
   // Not- Aus Taster Farbe 01 -- DB810.DBX67.5
   //    UN    "NA_SchrankFarbe"
   //    =      "DB820_Error_general".Machine[1].EmergencyStop.ColorUnit_01

   // Not- Aus Taster Farbe 02 -- DB810.DBX67.6
   //    UN    "NA_SchrankFarbe"
   //    =      "DB820_Error_general".Machine[1].EmergencyStop.ColorUnit_02

   // Not- Aus Taster an der Containerstation Komponente 1 wurde betätigt -- DB810.DBX67.1
   //    =     "DB820_Error_general".Machine[1].EmergencyStop.ContStation_C1
   // Not- Aus Taster an der Containerstation Komponente 2 wurde betätigt -- DB810.DBX67.2
   //    =     "DB820_Error_general".Machine[1].EmergencyStop.ContStation_C2

   // Not- Aus Signal von der Fremdanlage 1 steht an -- DB810.DBX67.3
         AN    "ES_Central";
         CLR;
         =     "DB820_Error_general".Machine[1].EmergencyStop.External_Plant_1;
   // Not- Aus  !! Reserve !!
         CLR;
         =     "DB820_Error_general".Machine[1].EmergencyStop.AdditionalComponent;
   // Not- Aus  !! Reserve !!
   //    =     "DB820_Error_general".Machine[1].EmergencyStop.Spare_1_5
   // Not- Aus  !! Reserve !!
   //    =      "DB820_Error_general".Machine[1].EmergencyStop.Spare_1_6

   // Not- Aus Taster an der Hydraulik Komponente 1 wurde betätigt -- DB810.DBX68.0
   //    =      "DB820_Error_general".Machine[1].EmergencyStop_Hydraulic[1]
   // Not- Aus Taster an der Hydraulik Komponente 2 wurde betätigt -- DB810.DBX68.1
   //    =      "DB820_Error_general".Machine[1].EmergencyStop_Hydraulic[2]
   // Not- Aus Taster an der Hydraulik Komponente 3 wurde betätigt -- DB810.DBX68.2
   //    =      "DB820_Error_general".Machine[1].EmergencyStop_Hydraulic[3]
   // Not- Aus Taster an der Hydraulik Komponente 4 wurde betätigt -- DB810.DBX68.3
   //    =      "DB820_Error_general".Machine[1].EmergencyStop_Hydraulic[4]
   // Not- Aus Taster an der Hydraulik Komponente 5 wurde betätigt -- DB810.DBX68.4
   //    =      "DB820_Error_general".Machine[1].EmergencyStop_Hydraulic[5]
   // Not- Aus Taster an der Hydraulik Komponente 6 wurde betätigt -- DB810.DBX68.5
   //    =      "DB820_Error_general".Machine[1].EmergencyStop_Hydraulic[6]
   // Not- Aus Taster an der Hydraulik Komponente 7 wurde betätigt -- DB810.DBX68.6
   //    =      "DB820_Error_general".Machine[1].EmergencyStop_Hydraulic[7]
   // Not- Aus Taster an der Hydraulik Komponente 8 wurde betätigt -- DB810.DBX68.7
   //    =      "DB820_Error_general".Machine[1].EmergencyStop_Hydraulic[8]

   //--------------------------------------------------------------------------------
   // Not- Aus Taster am Bedienpult Mischkopf 01 wurde betätigt
         A     "DB123_MH_IO_Signals".MH[1].IN.MH_EmergencyStop;
         =     "DB824_Error_MH_CP".EmergencyStop_Opanel_MH[1];
   //--------------------------------------------------------------------------------
   // Not- Aus Taster am Bedienpult Mischkopf 02 wurde betätigt
         A     "DB123_MH_IO_Signals".MH[2].IN.MH_EmergencyStop;
         =     "DB824_Error_MH_CP".EmergencyStop_Opanel_MH[2];
   //--------------------------------------------------------------------------------
   // Not- Aus Taster am Bedienpult Mischkopf 03 wurde betätigt
         A     "DB123_MH_IO_Signals".MH[3].IN.MH_EmergencyStop;
         =     "DB824_Error_MH_CP".EmergencyStop_Opanel_MH[3];
   //--------------------------------------------------------------------------------
   // Not- Aus Taster am Bedienpult Mischkopf 04 wurde betätigt
         A     "DB123_MH_IO_Signals".MH[4].IN.MH_EmergencyStop;
         =     "DB824_Error_MH_CP".EmergencyStop_Opanel_MH[4];
   //--------------------------------------------------------------------------------
   // Not- Aus Taster am Bedienpult Mischkopf 05 wurde betätigt
         A     "DB123_MH_IO_Signals".MH[5].IN.MH_EmergencyStop;
         =     "DB824_Error_MH_CP".EmergencyStop_Opanel_MH[5];
   //--------------------------------------------------------------------------------
   // Not- Aus Taster am Bedienpult Mischkopf 06 wurde betätigt
         A     "DB123_MH_IO_Signals".MH[6].IN.MH_EmergencyStop;
         =     "DB824_Error_MH_CP".EmergencyStop_Opanel_MH[6];
   //--------------------------------------------------------------------------------
   // Not- Aus Taster am Bedienpult Mischkopf 07 wurde betätigt
         A     "DB123_MH_IO_Signals".MH[7].IN.MH_EmergencyStop;
         =     "DB824_Error_MH_CP".EmergencyStop_Opanel_MH[7];
   //--------------------------------------------------------------------------------
   // Not- Aus Taster am Bedienpult Mischkopf 08 wurde betätigt
         A     "DB123_MH_IO_Signals".MH[8].IN.MH_EmergencyStop;
         =     "DB824_Error_MH_CP".EmergencyStop_Opanel_MH[8];
   //--------------------------------------------------------------------------------
   // Not- Aus Taster am Bedienpult Mischkopf 09 wurde betätigt
         A     "DB123_MH_IO_Signals".MH[9].IN.MH_EmergencyStop;
         =     "DB824_Error_MH_CP".EmergencyStop_Opanel_MH[9];
   //--------------------------------------------------------------------------------
   // Not- Aus Taster am Bedienpult Mischkopf 10 wurde betätigt
         A     "DB123_MH_IO_Signals".MH[10].IN.MH_EmergencyStop;
         =     "DB824_Error_MH_CP".EmergencyStop_Opanel_MH[10];
   //--------------------------------------------------------------------------------
   // Not- Aus Taster am Bedienpult Mischkopf 11 wurde betätigt
         A     "DB123_MH_IO_Signals".MH[11].IN.MH_EmergencyStop;
         =     "DB824_Error_MH_CP".EmergencyStop_Opanel_MH[11];
   //--------------------------------------------------------------------------------
   // Not- Aus Taster am Bedienpult Mischkopf 12 wurde betätigt
         A     "DB123_MH_IO_Signals".MH[12].IN.MH_EmergencyStop;
         =     "DB824_Error_MH_CP".EmergencyStop_Opanel_MH[12];
   //--------------------------------------------------------------------------------
   // Not- Aus Taster am Bedienpult Mischkopf 13 wurde betätigt
   //    =     "DB824_Error_MH_CP".Machine[1].EmergencyStop_Opanel_MH[13]
   // Not- Aus Taster am Bedienpult Mischkopf 14 wurde betätigt
   //    =     "DB824_Error_MH_CP".Machine[1].EmergencyStop_Opanel_MH[14]
   // Not- Aus Taster am Bedienpult Mischkopf 15 wurde betätigt
   //    =     "DB824_Error_MH_CP".Machine[1].EmergencyStop_Opanel_MH[15]
   // Not- Aus Taster am Bedienpult Mischkopf 16 wurde betätigt
   //    =     "DB824_Error_MH_CP".Machine[1].EmergencyStop_Opanel_MH[16]

   // Not- Aus Signal vom Formträger 01 steht an
         AN    "ES_MC01";
         CLR;
         =     "DB825_Error_Interface".EmergencyStop_MC[1];
   // Not- Aus Signal vom Formträger 02 steht an
         AN    "ES_MC02";
         CLR;
         =     "DB825_Error_Interface".EmergencyStop_MC[2];
   // Not- Aus Signal vom Formträger 03 steht an
         AN    "ES_MC03";
         CLR;
         =     "DB825_Error_Interface".EmergencyStop_MC[3];
   // Not- Aus Signal vom Formträger 04 steht an
         AN    "ES_MC04";
         CLR;
         =     "DB825_Error_Interface".EmergencyStop_MC[4];
   // Not- Aus Signal vom Formträger 05 steht an -- DB810.DBX72.4
   //    =      "DB820_Error_general".Machine[1].EmergencyStop_MC[5]
   // Not- Aus Signal vom Formträger 06 steht an -- DB810.DBX72.5
   //    =      "DB820_Error_general".Machine[1].Machine[1].EmergencyStop_MC[6]
   // Not- Aus Signal vom Formträger 07 steht an -- DB810.DBX72.6
   //    =      "DB820_Error_general".EmergencyStop_MC[7]
   // Not- Aus Signal vom Formträger 08 steht an -- DB810.DBX72.7
   //    =      "DB820_Error_general".Machine[1].EmergencyStop_MC[8]
   // Not- Aus Signal vom Formträger 09 steht an -- DB810.DBX73.0
   //    =      "DB820_Error_general".Machine[1].EmergencyStop_MC[9]
   // Not- Aus Signal vom Formträger 10 steht an -- DB810.DBX73.1
   //    =      "DB820_Error_general".Machine[1].EmergencyStop_MC[10]
   // Not- Aus Signal vom Formträger 11 steht an -- DB810.DBX73.2
   //    =      "DB820_Error_general".Machine[1].EmergencyStop_MC[11]
   // Not- Aus Signal vom Formträger 12 steht an -- DB810.DBX73.3
   //    =      "DB820_Error_general".Machine[1].EmergencyStop_MC[12]
   // Not- Aus Signal vom Formträger 13 steht an -- DB810.DBX73.4
   //    =      "DB820_Error_general".Machine[1].EmergencyStop_MC[13]
   // Not- Aus Signal vom Formträger 14 steht an -- DB810.DBX73.5
   //    =      "DB820_Error_general".Machine[1].Machine[1].EmergencyStop_MC[14]
   // Not- Aus Signal vom Formträger 15 steht an -- DB810.DBX73.6
   //    =      "DB820_Error_general".EmergencyStop_MC[15]
   // Not- Aus Signal vom Formträger 16 steht an -- DB810.DBX73.7
   //    =      "DB820_Error_general".Machine[1].EmergencyStop_MC[16]
   // Automatik- Stop Schutztür zum Roboterbereich 1 steht noch an -- DB810.DBX74.0
   //    U     "ES_SaftyDoorRobot"
   //    =     "DB820_Error_general".Machine[1].Safety_Door_selected[1]
   // Automatik- Stop Schutztür zum Roboterbereich 2 steht noch an -- DB810.DBX74.1
   //    =      "DB820_Error_general".Machine[1].Safty_Door_selected[2]
   // Automatik- Stop Schutztür zum Rovingbereich 1 steht noch an -- DB810.DBX74.2
   //    =      "DB820_Error_general".Machine[1].Safty_Door_selected[3]
   // Automatik- Stop Schutztür zum Rovingbereich 2 steht noch an -- DB810.DBX74.3
   //    =      "DB820_Error_general".Machine[1].Safty_Door_selected[4]
   // Die Vorwahl zum öffnen der Schutztür Roving 1 aktiv -- DB810.DBX74.4
   //    =      "DB820_Error_general".Machine[1].Safty_Door_selected[5]
   // Die Vorwahl zum öffnen der Schutztür Roving 2 aktiv -- DB810.DBX74.5
   //    =      "DB820_Error_general".Machine[1].Safty_Door_selected[6]
   // Die Vorwahl zum öffnen der Schutztür Roboter 1 aktiv -- DB810.DBX74.6
   //    =      "DB820_Error_general".Machine[1].Safty_Door_selected[7]
   // Die Vorwahl zum öffnen der Schutztür Roboter 2 aktiv -- DB810.DBX74.7
   //    =      "DB820_Error_general".Machine[1].Safty_Door_selected[8]
   // Betriebsart Testen  ist angewählt  -- DB820.DBX62.0
         A     "DB619_State_MPart".Operationmode[1].Test;
         =     "DB820_Error_general".Machine[1].OpMode_Test;
   // Wochenendschaltung Maschine 1  -- DB810.DBX76.1
   //-----------------------------------------------------------------------
         A     "DB619_State_MPart".Recirculation[1].Weekendswitching;
         A     "DB619_State_MPart".Recirculation[1].Switch_Reduced;
         AN    "DB009_Faults".Fault_State_Grp_1_M1;
         =     "DB820_Error_general".Machine[1].Weekend_Mode;
   // Wochenendschaltung Maschine 2  -- DB810.DBX94.1
   //------------------------------------------------------------------------
         A     "DB619_State_MPart".Recirculation[2].Weekendswitching;
         A     "DB619_State_MPart".Recirculation[2].Switch_Reduced;
         AN    "DB009_Faults".Fault_State_Grp_1_M2;
         =     "DB820_Error_general".Machine[2].Weekend_Mode;
   // Automatik- Stop ist noch nicht quittiert -- DB810.DBX76.4
         AN    "AS";
         CLR;
         =     "DB820_Error_general".Machine[1].AutoStop;
END_REGION

REGION Network 6: Additional bits for emergency stop
   // Emergency stop machine poly 1
   //    U     "ES_K1"
   //    =     "DB820_Error_general".Machine[1].EmergencyStop[1]

   // Emergency stop machine poly 2
   //    U     "ES_K2"
   //    =     "DB820_Error_general".Machine[1].EmergencyStop[2]

   // Emergency stop machine poly 3
   //    U     "ES_K3"
   //    =     "DB820_Error_general".Machine[1].EmergencyStop[3]

   // Emergency stop machine poly 4
   //    U     "ES_K4"
   //    =     "DB820_Error_general".Machine[1].EmergencyStop[4]

   // Emergency stop machine iso 1
   //    U     "ES_K5"
   //    =     "DB820_Error_general".Machine[1].EmergencyStop[5]

   // Emergency stop machine iso 2
   //    U     "ES_K6"
   //    =     "DB820_Error_general".Machine[1].EmergencyStop[6]

   // Emergency stop main cabinet
   //    U     "ES_ctrl_cabinet_conveyor"
   //    =     "DB820_Error_general".Machine[1].EmergencyStop[7]

   // Emergency stop operating panel of conveyor
   //    U     "ES_OP_handlingarea"
   //    =     "DB820_Error_general".Machine[1].EmergencyStop[8]

   // Emergency stop safety door toolchange
   //    U     "ES_op_changing_unit"
   //    =     "DB820_Error_general".Machine[1].EmergencyStop[9]

   // Emergency stop safety door chain tensioner
   //    U     "ES_door_Entr_Conveyor"
   //    =     "DB820_Error_general".Machine[1].EmergencyStop[10]

   // Emergency stop safety door to robot 1
   //    U     "ES_door_robot_MH1"
   //    =     "DB820_Error_general".Machine[1].EmergencyStop[11]

   // Emergency stop safety door to robot 2
   //    U     "ES_door_robot_MH2"
   //    =     "DB820_Error_general".Machine[1].EmergencyStop[12]

   // Emergency stop mushroom picking
   //    U     "ES_mushroom_picking"
   //    =     "DB820_Error_general".Machine[1].EmergencyStop[13]

   // Emergency stop chain monitoring
   //    U     "ES_chain_tight"
   //    =     "DB820_Error_general".Machine[1].EmergencyStop[14]
END_REGION
END_FUNCTION

FUNCTION "FC082_FaultProfiBus" : Void   // FC82, STL
TITLE = Faults at profibus net
{ S7_Optimized_Access := 'FALSE' }
VERSION : 0.1
   VAR_TEMP
      Null : Byte;
      ERROR_CODE : Int;
   END_VAR
BEGIN

REGION Network 1: Rücksetzen Störungen Profibus Maschine 1
         A     "DB009_Faults".Faults_Reset_FKT_M1;
         JCN   nres;

         L     0;
         T     #Null;

         CALL  FILL
         ( BVAL    := #Null,
           RET_VAL := #ERROR_CODE,
           BLK     := "DB820_Error_general".Profibus_DP[1]
         );

   nres: NOP   0;
END_REGION

REGION Network 2: Störungsauswertung Profibus Maschine 1
   // Profinet-IO
   // ProNet Modul 01 machine not available on profinet
         A     "PN_AI".Module[1].AI8.Active;
         A     "PN_AI".Module[1].AI8.ChckConnFault;
         ON    "PN_Devices".Device_available[1];
         AN    "DB820_Error_general".Profibus_DP[1].Member[1];
         S     "DB009_Faults".Faultschanging_M1;
         S     "DB009_Faults".Faults_FKT_Grp_3_M1;
         S     "DB820_Error_general".Profibus_DP[1].Member[1];


   // ProNet Modul 02 mixing head not available on profinet
         A     "PN_AI".Module[2].AI8.Active;
         A     "PN_AI".Module[2].AI8.ChckConnFault;
         ON    "PN_Devices".Device_available[2];
         AN    "DB820_Error_general".Profibus_DP[1].Member[2];
         S     "DB009_Faults".Faultschanging_M1;
         S     "DB009_Faults".Faults_FKT_Grp_3_M1;
         S     "DB820_Error_general".Profibus_DP[1].Member[2];


   // pn-pn coupler not available on profinet
         ON    "PN_Devices".Device_available[3];
         AN    "DB820_Error_general".Profibus_DP[1].Member[3];
         CLR;
         S     "DB009_Faults".Faultschanging_M1;
         S     "DB009_Faults".Faults_FKT_Grp_3_M1;
         S     "DB820_Error_general".Profibus_DP[1].Member[3];
END_REGION
END_FUNCTION

FUNCTION "FC089_quit_Faults" : Void   // FC89, STL
TITLE = Confirme faults machine 1..4 and plants
{ S7_Optimized_Access := 'FALSE' }
AUTHOR : KT242
FAMILY : RS_KK
NAME : Fault_oK
VERSION : 1.1
// Die Stoerungsquittierung erfolgt in zwei SPS-Zyklen: 
// 1.: mit Reset_fault_Fkt werden die Störungsbits der einzelnen FCs zurückgesetzt
// 2.: mit Reset_fault_Grp werden die Störungsbits der FCs für die Störungsgruppen
//     zurückgesetzt. Bilden diese nun die Störungen neu, so werten sie von
//     den einzelnen FCs bereits den aktuellen Stand aus, da diese bereits einen
//     SPS-Zyklus früher bearbeitet wurden.
// 
// Das Ablöschen der Störungsbits an die Visualisierung wird von den einzelnen 
// Stör-FCs organisiert.
   VAR_INPUT
      IN_Button_Acknowledge : Bool;   // Button to acknowledge malfunctions (quit)
      IN_Button_Horn_Off : Bool;   // Button to switch off the Horn
      IN_First_PLC_cycle : Bool;   // Pulse start up PLC to erase faults
      IN_IndicatorLampTest : Bool;   // Button to test indicator lamps
      IN_Fault_Grp_1_active_M1 : Bool;   // Fault flag of active fault level 1 of machine 1
      IN_Fault_Grp_2_active_M1 : Bool;   // Fault flag of active fault level 2 of machine 1
      IN_Fault_Grp_3_active_M1 : Bool;   // Fault flag of active fault level 3 of machine 1
      IN_Fault_Grp_1_active_M2 : Bool;   // Fault flag of active fault level 1 of machine 2
      IN_Fault_Grp_2_active_M2 : Bool;   // Fault flag of active fault level 2 of machine 2
      IN_Fault_Grp_3_active_M2 : Bool;   // Fault flag of active fault level 3 of machine 2
      IN_Fault_Grp_1_active_M3 : Bool;   // Fault flag of active fault level 1 of machine 3
      IN_Fault_Grp_2_active_M3 : Bool;   // Fault flag of active fault level 2 of machine 3
      IN_Fault_Grp_3_active_M3 : Bool;   // Fault flag of active fault level 3 of machine 3
      IN_Fault_Grp_1_active_M4 : Bool;   // Fault flag of active fault level 1 of machine 4
      IN_Fault_Grp_2_active_M4 : Bool;   // Fault flag of active fault level 2 of machine 4
      IN_Fault_Grp_3_active_M4 : Bool;   // Fault flag of active fault level 3 of machine 4
      IN_Fault_Grp_1_active_AP : Bool;   // Fault flag of active fault level 1 of external plant
      IN_Fault_Grp_2_active_AP : Bool;   // Fault flag of active fault level 2 of external plant
      IN_Fault_Grp_3_active_AP : Bool;   // Fault flag of active fault level 3 of external plant
   END_VAR
   VAR_OUTPUT
      OUT_acoustical_indicator : Bool;   // Ausgang für eine akustische Störungsanzeige (Nur bei Neustörungen)
      OUT_optical_indicator : Bool;   // Ausgang für eine optische Störungsanzeige
   END_VAR
   VAR_IN_OUT
      IO_Fault_changed_M1 : Bool;   // Feststellen einer Störungsänderung of machine 1 für Abarbeitung
      IO_Fault_changed_M2 : Bool;   // Feststellen einer Störungsänderung of machine 2 für Abarbeitung
      IO_Fault_changed_M3 : Bool;   // Feststellen einer Störungsänderung of machine 3 für Abarbeitung
      IO_Fault_changed_M4 : Bool;   // Feststellen einer Störungsänderung of machine 4 für Abarbeitung
      IO_Fault_changed_AP : Bool;   // Feststellen einer Störungsänderung von der Fremdanlage für Abarbeitung
      IO_Horn : Bool;   // Hilfsmerker zum ablöschen der akustischen Störanzeige nach Quittierung
      IO_Reset_fault_Grp : Bool;   // Signal zum quittieren der Störungen innerhalb der Störungsbausteine
      IO_Reset_fault_Fkt : Bool;   // Signal zum quittieren der Störungen innerhalb der einzelnen Funktionsbausteine
      IO_Quit_Edge : Bool;   // Hilkfsmerker zur Überwachung der Betätigung des Quittiertasters
   END_VAR
   VAR_TEMP
      Overall_Fault_Flag : Bool;   // Zwischenmerker für die erkennung einer anliegenden Störung
      Quit_Flanke : Bool;   // Zwischenmerker als Impuls für die Störungsquittierung
      New_Fault : Bool;
   END_VAR
BEGIN

REGION Network 1: Acknowledge (quit) faults of fault levels at PLC
   // Über das Bit Reset_fault_Fkt werden zuerst die Störungen in den Funktionen in 
   // dem sie gebildet werden abgelöscht. Im nächsten SPS- Zyklus werden dann erst 
   // die Störbits in den jeweiligen Störungsbausteinen abgelöscht
         A     #IO_Reset_fault_Grp;  // Für den Störungsbaustein
         R     #IO_Reset_fault_Grp;
         A     #IO_Reset_fault_Fkt;  // Für die einzelnen Funktionsbausteine
         S     #IO_Reset_fault_Grp;
         A     #IO_Reset_fault_Grp;
         R     #IO_Reset_fault_Fkt;
END_REGION

REGION Network 2: Bilden einer Sammelstörung
   // Für die Erkennung der Störungsänderung wird eine Sammelstörung benötigt. 
   // Diese wird aus allen eingehenden Störungen gebildet.
         O     #IN_Fault_Grp_1_active_M1;
         O     #IN_Fault_Grp_2_active_M1;
         O     #IN_Fault_Grp_3_active_M1;
         O     #IN_Fault_Grp_1_active_M2;
         O     #IN_Fault_Grp_2_active_M2;
         O     #IN_Fault_Grp_3_active_M2;
         O     #IN_Fault_Grp_1_active_M3;
         O     #IN_Fault_Grp_2_active_M3;
         O     #IN_Fault_Grp_3_active_M3;
         O     #IN_Fault_Grp_1_active_M4;
         O     #IN_Fault_Grp_2_active_M4;
         O     #IN_Fault_Grp_3_active_M4;
         O     #IN_Fault_Grp_1_active_AP;
         O     #IN_Fault_Grp_2_active_AP;
         O     #IN_Fault_Grp_3_active_AP;
         =     #Overall_Fault_Flag;
END_REGION

REGION Network 3: Quittierflanke gegen Dauerbetätigung des Quittiertasters
   // Damit zum quittieren der Störungen bewußt der Taster zwei betätigt werden muß 
   // wird hier die Änderung des Quittiertasters für das Programm verwendet.
         O     #IN_Button_Acknowledge;
         FP    #IO_Quit_Edge;
         =     #Quit_Flanke;
END_REGION

REGION Network 4: Hilfsmerker für die Störungsbildung zurücksetzen
   // Wenn keine Störung mehr ansteht oder
   // Wenn eine neue Störungsänderung erfolgt,
   // wird das Bit für die erste Quittierung zurückgesetzt
         O     #IO_Fault_changed_M1;
         O     #IO_Fault_changed_M2;
         O     #IO_Fault_changed_M3;
         O     #IO_Fault_changed_M4;
         O     #IO_Fault_changed_AP;
         ON    #Overall_Fault_Flag;
         R     #IO_Horn;
END_REGION

REGION Network 5: Quittierbit für die Störbits innerhalb der einzelnen Funktionen
   // Das Bit zum ablöschen der Störungsbits innerhalb der einzelnen 
   // Funktionsbausteinen, welches auch gleichzeitig das Quittierbit an die 
   // Visualisierung ist, wird gesetzt, wenn:
   // - Wenn Störungen anstehen und zum 2´ten mal quittiert wird, 
   // - Keine Störungen anstehen und der Quittiertsater betätigt wird und
   // - Beim einschalten der Steuerung.
         A     #Overall_Fault_Flag;
         A     #IO_Horn;
         A     #Quit_Flanke;
         O;
   //
         AN    #Overall_Fault_Flag;
         A     #IN_Button_Acknowledge;
   //
         O     #IN_First_PLC_cycle;
         S     #IO_Reset_fault_Fkt;
END_REGION

REGION Network 6: Rücksetzen des Bits für die Erste Quittierung
   // Diese Bit wird benötigt, um die akustische Störungsanzeige nach der ersten 
   // Quittierung auszuschalten. Aber auch für die allgemeine Erkennung des erneuten 
   // betätigen des Quittiertasters.
   // Wurde das Quittierbit für die einzelnen Maschinen gesetzt, wird das Bit 
   // für für die 1´te Quittierung zurückgesetzt
         A     #IO_Reset_fault_Fkt;
         R     #IO_Horn;
   //
         A     #Overall_Fault_Flag;
         A     #Quit_Flanke;
         O     #IN_Button_Horn_Off;
         AN    #IO_Reset_fault_Fkt;
         AN    #IO_Fault_changed_M1;
         AN    #IO_Fault_changed_M2;
         AN    #IO_Fault_changed_M3;
         AN    #IO_Fault_changed_AP;
         S     #IO_Horn;
END_REGION

REGION Network 7: Ansteuern der optischen Störungsanzeige
   // Die optische Anzeige der Störung wird immer angesteuert, solange eine Störung 
   // vorhanden ist, oder wenn die Funktion "Lampentest" aktiv ist.
         A     #Overall_Fault_Flag;
         A     "Flag_01_000_Hertz";
         O     #IN_IndicatorLampTest;
         =     #OUT_optical_indicator;
END_REGION

REGION Network 8: Ansteuern der akustischen Störungsanzeige
   // Die akustische Störungsanzeige wird nur angesteuert, bis die erste Quittierung 
   // über den Quittiertaster erfolgte. 
   // Sobald eine neue Störung erkannt wurde, oder die Störung nach dem erneuten 
   // betätigen des Quittiertasters noch immer ansteht wird die akustische 
   // Störungsanzeige erneut aktiv.
         A     #Overall_Fault_Flag;
         A     "Flag_01_000_Hertz";
         AN    #IO_Horn;
         =     #OUT_acoustical_indicator;
END_REGION

REGION Network 9: Rücksetzen der Störungsänderungen
   // Die Bits für die Information einer Störungsänderung aus den Störungsbausteinen 
   // der Maschinen oder der Anlage wird zurückgesetzt. Hierdurch kann bei einer 
   // Neustörung dieses Bit wieder neu gestzt werden.
         AN    #IN_First_PLC_cycle;
         R     #IO_Fault_changed_M1;
         R     #IO_Fault_changed_M2;
         R     #IO_Fault_changed_M3;
         R     #IO_Fault_changed_M4;
         R     #IO_Fault_changed_AP;
END_REGION
END_FUNCTION

FUNCTION "FC091_PouringCycle" : Void   // FC91, STL
TITLE = Shot cycle
{ S7_Optimized_Access := 'FALSE' }
AUTHOR : KT242
FAMILY : RS_KK
NAME : PCycle
VERSION : 1.3
// The function organizes the sequence of a shot cycle.
// With the start shot signal the following happens: 
// 1a: when no cycle is active the Pressurize Time starts
// 1b: when the StandByTime is active the CntrlChangeTime starts
// 2: after PressurizeTime or CntrlCnangeTime the shot is enabled
// 4. after the shot the StandByTime is started
// 5. if during the StandByTime no new cycle ist started, the cycle is finished.
   VAR_INPUT
      IN_OMAutomatic : Bool;   // Foaming machine in automatic mode
      IN_OMChange : Bool;   // Operation mode changed between service and shot with foam
      IN_ResetFaults : Bool;   // Bit to reset fault bits
      IN_LampTest : Bool;   // Lamptest activated
      IN_EnableCycle : Bool;   // External enable signal for shot cycle
      IN_EnablePressurizeTime : Bool;   // Release to start pressurize time (e.g. all pistons ready at KK machine)
      IN_ShotActive : Bool;   // Signal from ProCan module that shot is active
      IN_Hydraulics_OK : Bool;   // Pressure of hydraulic system is ok
      IN_DW_PressurizeTime : S5Time;   // Time for pressure build up with new start
      IN_DW_StandByTime : S5Time;   // Standby time for waiting for new shot start
      IN_DW_CntrlChangeTime : S5Time;   // Time between shots for changing controller values (flow, pressure,...)
      IN_DW_MaxWaitTime : S5Time;   // Timevalue for maximum waiting time for shot
      IN_DW_MaxShotTime : S5Time;   // Maximum value for shot
      IN_Cycletimer : Timer;   // Timer for internal use
      IN_FaultLevel_1 : Bool;
      IN_FaultLevel_2 : Bool;
   END_VAR
   VAR_OUTPUT
      OUT_LampMachineOK : Bool;   // Lamp machine is ready for foaming
   END_VAR
   VAR_IN_OUT
      IO_Status : ANY;   // Pointer to status signals for the shot cycle
      IO_Fault : ANY;
      IO_FaultLevel_1 : Bool;   // Fault message of level 1 is active and was not acknowledged
      IO_FaultLevel_2 : Bool;   // Fault message of level 2 is active and was not acknowledged
      IO_FaultLevel_3 : Bool;   // Fault message of level 3 is active and was not acknowledged
      IO_NewFault : Bool;
      IO_StartShotCycle : Bool;   // Start signal for shot cycle
      IO_StopShotCycle : Bool;   // Stop signal for shot cycle
   END_VAR
   VAR_TEMP
      Temp_IO_Status : "UDT091_PouringCycleState";   // Temporary informations for the shot cycle
      Temp_IO_Fault : "UDT1819_FLT_PouringCycle";   // Fault bits for the shot cycle
      ERROR_CODE : Int;   // Error state of systemfunction "BLKMOV" Blockmove
      AnyPointer1 : ANY;   // Pointer to copy thr array "IO_Status" and "Temp_IO_Status"
      AnyPointer2 : ANY;   // Pointer to copy thr array "IO_Status" and "Temp_IO_Status"
      TimeValue : Time;   // Variable for calculation of time for pressure request to hydraulic
      TimeValueS5Time : S5Time;
   END_VAR
BEGIN

REGION Network 1: Saved data integration
   //-----
         L;
         LAR1;
         LAR2;
   //-----
         L     W[AR1, P#0.0];  // Bytes
         T     W[AR2, P#0.0];
         L     W[AR1, P#2.0];  // Amount of bytes
         T     W[AR2, P#2.0];
         L     W[AR1, P#4.0];  // Block no,
         T     W[AR2, P#4.0];
         L     D[AR1, P#6.0];  // Startadress of data
         T     D[AR2, P#6.0];
   //-----
         CALL  BLKMOV
         ( SRCBLK  := #AnyPointer1,
           RET_VAL := #ERROR_CODE,
           DSTBLK  := #Temp_IO_Status
         );
   //-----
         L;
         LAR1;
         LAR2;
   //-----
         L     W[AR1, P#0.0];  // Bytes
         T     W[AR2, P#0.0];
         L     W[AR1, P#2.0];  // Amount of bytes
         T     W[AR2, P#2.0];
         L     W[AR1, P#4.0];  // Block no,
         T     W[AR2, P#4.0];
         L     D[AR1, P#6.0];  // Startadress of data
         T     D[AR2, P#6.0];
   //-----
         CALL  BLKMOV
         ( SRCBLK  := #AnyPointer2,
           RET_VAL := #ERROR_CODE,
           DSTBLK  := #Temp_IO_Fault
         );
   //-----
END_REGION

REGION Network 2: Reset Faults
   //-----
         A     #IN_ResetFaults;
         R     #Temp_IO_Fault.FLT_KLZ_0;
         R     #Temp_IO_Fault.FLT_OP_Mode;
         R     #Temp_IO_Fault.FLT_Max_Shottime;
         R     #Temp_IO_Fault.FLT_Max_Waittime;
   //-----
END_REGION

REGION Network 3: Enable cycle
         O(;
         L     #IN_DW_PressurizeTime;
         L     0;
         ==I;
         );
         O(;
         L     #IN_DW_StandByTime;
         L     0;
         ==I;
         );
         O(;
         L     #IN_DW_CntrlChangeTime;
         L     0;
         ==I;
         );
         O(;
         L     #IN_DW_MaxWaitTime;
         L     0;
         ==I;
         );
         O(;
         L     #IN_DW_MaxShotTime;
         L     0;
         ==I;
         );
         AN    #Temp_IO_Fault.FLT_KLZ_0;
         S     #Temp_IO_Fault.FLT_KLZ_0;  // Störung Zeit nicht programmiert
         S     #IO_NewFault;
   //
         ON    #IN_FaultLevel_2;
         O     #Temp_IO_Status.running;
         AN    #IN_FaultLevel_1;
         A     #IN_OMAutomatic;
         A     #IN_Hydraulics_OK;
         AN    #Temp_IO_Fault.FLT_KLZ_0;
         A     #IN_EnableCycle;
         =     #Temp_IO_Status.Release;
END_REGION

REGION Network 4: Finish cycle
   //--------------------------------------------------------------------
   // 4. Reset signals at cycle end
   //--------------------------------------------------------------------
         A     #Temp_IO_Status.PulseCycleEnd;
         R     #Temp_IO_Status.running;
         R     #Temp_IO_Status.PulseCycleEnd;
         R     #Temp_IO_Status.MHWasOpen;
         R     #Temp_IO_Status.CtrlChangeTimeRuns;
         R     #Temp_IO_Status.PulsShotend;
         R     #Temp_IO_Status.ShotRuns;
         R     #Temp_IO_Status.StandByTimeRuns;
   //--------------------------------------------------------------------
   // 1. Finish foamingcycle recirculation not necessary
   //--------------------------------------------------------------------
         O(;
         O     #IO_StopShotCycle;
         AN    #Temp_IO_Status.MHWasOpen;
         );
         O     #IN_FaultLevel_1;
         ON    #Temp_IO_Status.Release;
         O     #Temp_IO_Status.RmpStandByTimeEnd;
         O     #Temp_IO_Fault.FLT_Max_Waittime;
         S     #Temp_IO_Status.PulseCycleEnd;
         R     #Temp_IO_Status.PressurizeTimeFinished;
   //--------------------------------------------------------------------
   // 3. Finish foamingcycle during changetime -> recirculation necessary
   //--------------------------------------------------------------------
         O     #IN_FaultLevel_1;
         O     #IO_StopShotCycle;
         ON    #Temp_IO_Status.Release;
         A(;
         O(;
         A     #Temp_IO_Status.PressurizeTimeFinished;
         A     #Temp_IO_Status.MHWasOpen;
         );
         O     #Temp_IO_Status.CtrlChangeTimeRuns;
         );
         S     #Temp_IO_Status.StandByTimeRuns;
         R     #Temp_IO_Status.CtrlChangeTimeRuns;
         R     #Temp_IO_Status.MHWasOpen;
   //------------------------------------------------------------------
   // 2. Finish foamingcycle recirculation necessary
   //------------------------------------------------------------------
         A     #Temp_IO_Status.Release;
         AN    #Temp_IO_Status.PulseCycleEnd;
         AN    #Temp_IO_Fault.FLT_Max_Shottime;
         AN    #IO_StopShotCycle;
         AN    #IN_FaultLevel_1;
         JC    actv;
   //-----
         R     #Temp_IO_Status.PressurizeTimeRuns;
         R     #Temp_IO_Status.RmpPressurizeTimeEnd;
         R     #Temp_IO_Status.RmpStandByTimeEnd;
         R     #Temp_IO_Status.RmpCtrlChangeTimeEnd;
         R     #Temp_IO_Status.Shotrelease;
         R     #Temp_IO_Status.SelectHydForShot;
   //-----
         CLR;
         L     S5T#0MS;
         SP    #IN_Cycletimer;
         JU    save;
   //-----
   actv: NOP   0;
   //-----
END_REGION

REGION Network 5: Start cycle if no cycle is active
   //-----
         AN    #IO_StartShotCycle;
         JC    nosr;
   //-----
         R     #IO_StartShotCycle;
   //-----
         A     #Temp_IO_Status.StandByTimeRuns;
         R     #Temp_IO_Status.StandByTimeRuns;
         R     #Temp_IO_Status.RmpStandByTimeEnd;
         S     #Temp_IO_Status.CtrlChangeTimeRuns;
         JCN   strc;
   //-----
         CLR;
         L     S5T#0MS;
         SP    #IN_Cycletimer;
   //-----
   strc: AN    #Temp_IO_Status.running;
         S     #Temp_IO_Status.running;
   //-----
   nosr: NOP   0;
   //-----
END_REGION

REGION Network 6: Pressurize time
   //-----
         O     #Temp_IO_Status.PressurizeTimeFinished;
         ON    #Temp_IO_Status.running;
         O     #Temp_IO_Status.MHWasOpen;
         JC    pten;
   //-----
         A     #Temp_IO_Status.PressurizeTimeRuns;
         AN    #Temp_IO_Status.RmpPressurizeTimeEnd;
         L     #IN_DW_PressurizeTime;
         SD    #IN_Cycletimer;
   //-----
         A     #IN_EnablePressurizeTime;
         S     #Temp_IO_Status.PressurizeTimeRuns;
   //-----
         A     #Temp_IO_Status.RmpPressurizeTimeEnd;
         R     #Temp_IO_Status.RmpPressurizeTimeEnd;
         R     #Temp_IO_Status.PressurizeTimeRuns;
         S     #Temp_IO_Status.PressurizeTimeFinished;
         S     #Temp_IO_Status.Shotrelease;
   //-----
         A     #IN_Cycletimer;
         S     #Temp_IO_Status.RmpPressurizeTimeEnd;
   //-----
   pten: NOP   0;
   //-----
END_REGION

REGION Network 7: Request hydraulic pressure before 1st shot
   //-----
         ON    #Temp_IO_Status.PressurizeTimeRuns;
         O     #Temp_IO_Status.SelectHydForShot;
         JC    nhyd;
   //-----
         LC    #IN_Cycletimer;
         T     #TimeValueS5Time;
         CALL  T_CONV
         ( IN  := #TimeValueS5Time,
           OUT := #TimeValue
         );
   //-----
         L     #TimeValue;
         L     2000;
         <D;
         S     #Temp_IO_Status.SelectHydForShot;
   //-----
   nhyd: NOP   0;
   //-----
END_REGION

REGION Network 8: Control change time
   //-----
         AN    #Temp_IO_Status.CtrlChangeTimeRuns;
         JC    ncct;
   //-----
         AN    #Temp_IO_Status.RmpCtrlChangeTimeEnd;
         L     #IN_DW_CntrlChangeTime;
         SD    #IN_Cycletimer;
   //-----
         A     #Temp_IO_Status.RmpCtrlChangeTimeEnd;
         R     #Temp_IO_Status.RmpCtrlChangeTimeEnd;
         R     #Temp_IO_Status.CtrlChangeTimeRuns;
         S     #Temp_IO_Status.Shotrelease;
   //-----
         A     #IN_Cycletimer;
         S     #Temp_IO_Status.RmpCtrlChangeTimeEnd;
   //-----
   ncct: NOP   0;
   //-----
END_REGION

REGION Network 9: Wait for shot
   //-----
         ON    #Temp_IO_Status.Shotrelease;
         JC    nrel;
         A     #IN_ShotActive;
         S     #Temp_IO_Status.ShotRuns;
   //-----
         A     #Temp_IO_Status.ShotRuns;
         JC    rt09;
   //-----
         A     #Temp_IO_Status.Shotrelease;
         L     #IN_DW_MaxWaitTime;
         SD    #IN_Cycletimer;
         A     #IN_Cycletimer;
         R     #Temp_IO_Status.Shotrelease;
   //-----
         A     #IN_Cycletimer;
         AN    #Temp_IO_Fault.FLT_Max_Waittime;
         S     #Temp_IO_Fault.FLT_Max_Waittime;
         S     #IO_NewFault;
   //-----
   rt09: ON    #Temp_IO_Status.ShotRuns;
         O     #Temp_IO_Status.MHWasOpen;
         AN    #Temp_IO_Fault.FLT_Max_Waittime;
         JC    nrel;
         CLR;
         L     S5T#0MS;
         SP    #IN_Cycletimer;
   //-----
   nrel: A     #IN_ShotActive;
         A     #Temp_IO_Status.Shotrelease;
         S     #Temp_IO_Status.MHWasOpen;
   //-----
END_REGION

REGION Network 10: Shot
   //-----
         A     #Temp_IO_Status.PulsShotend;
         R     #Temp_IO_Status.PulsShotend;
         R     #Temp_IO_Status.ShotRuns;
   //-----
         AN    #Temp_IO_Status.ShotRuns;
         JC    nsht;
         A     #IN_ShotActive;
         L     #IN_DW_MaxShotTime;
         SD    #IN_Cycletimer;
         A     #IN_Cycletimer;
         AN    #Temp_IO_Fault.FLT_Max_Shottime;
         S     #Temp_IO_Fault.FLT_Max_Shottime;
         S     #IO_NewFault;
   //-----
         ON    #IN_ShotActive;
         ON    #Temp_IO_Status.Shotrelease;
         A     #Temp_IO_Status.ShotRuns;
         S     #Temp_IO_Status.PulsShotend;
         NOP   0;
         S     #Temp_IO_Status.StandByTimeRuns;
         R     #Temp_IO_Status.Shotrelease;
   //-----
         AN    #Temp_IO_Status.PulsShotend;
         JC    nsht;
         CLR;
         L     S5T#0MS;
         SP    #IN_Cycletimer;
   //-----
   nsht: NOP   0;
   //-----
END_REGION

REGION Network 11: Stand by time
   //-----
         AN    #Temp_IO_Status.StandByTimeRuns;
         JC    nstb;
         AN    #Temp_IO_Status.RmpStandByTimeEnd;
         L     #IN_DW_StandByTime;
         SD    #IN_Cycletimer;
   //-----
         A     #Temp_IO_Status.RmpStandByTimeEnd;
         R     #Temp_IO_Status.RmpStandByTimeEnd;
         R     #Temp_IO_Status.StandByTimeRuns;
   //-----
         A     #IN_Cycletimer;
         S     #Temp_IO_Status.RmpStandByTimeEnd;
   //-----
   nstb: NOP   0;
   //-----
END_REGION

REGION Network 12: Lamp ready for operation
   //-----
   save: A     #Temp_IO_Status.Release;
         AN    #Temp_IO_Status.running;
         O;
         A     #Temp_IO_Status.running;
         AN    #Temp_IO_Status.ShotRuns;
         A     "Flag_01_000_Hertz";
         O;
         A     #Temp_IO_Status.ShotRuns;
         A     "Flag_05_000_Hertz";
         O     #IN_LampTest;
         =     #OUT_LampMachineOK;
   //-----
END_REGION

REGION Network 13: Error handling
   //-----
         A     #Temp_IO_Status.running;
         A     #Temp_IO_Status.ShotRuns;
         A     #IN_OMChange;
         AN    #Temp_IO_Fault.FLT_OP_Mode;
         S     #Temp_IO_Fault.FLT_OP_Mode;
         S     #IO_NewFault;
   //-----
         O     #Temp_IO_Fault.FLT_Max_Shottime;
         O     #Temp_IO_Fault.FLT_OP_Mode;
         S     #IO_FaultLevel_1;
   //-----
   //      O     XXXXXXXX
   //      S     #IO_FaultLevel_2
   //-----
         O     #Temp_IO_Fault.FLT_Max_Waittime;
         O     #Temp_IO_Fault.FLT_KLZ_0;
         S     #IO_FaultLevel_3;
   //-----
END_REGION

REGION Network 14: Save data
   //-----
         CALL  BLKMOV
         ( SRCBLK  := #Temp_IO_Status,
           RET_VAL := #ERROR_CODE,
           DSTBLK  := #AnyPointer1
         );
   //-----
         CALL  BLKMOV
         ( SRCBLK  := #Temp_IO_Fault,
           RET_VAL := #ERROR_CODE,
           DSTBLK  := #AnyPointer2
         );
   //-----
END_REGION
END_FUNCTION

FUNCTION "FC096_Faults_MH" : Void   // FC96, STL
TITLE = Faults of mixinghead during shot cycle
{ S7_Optimized_Access := 'FALSE' }
NAME : Faults
VERSION : 0.1
   VAR_INPUT
      IN_ProCanMH_State : Struct
         NoShotReleaseFromCP : Bool;   // No Shot Release from Cleaning Piston
         NoShotReleaseFromExtern : Bool;   // No Shot Release from Extern
         Ready4Shot : Bool;   // Ready for Shot
         shotactive_MH : Bool;   // Shot is active
         shotdone_MH : Bool;   // Shot finished
         Spare5 : Bool;
         Spare6 : Bool;
         Spare7 : Bool;
         SPFopening_MH : Bool;   // Steering piston fault opening time exceeded
         SPFclosing_MH : Bool;   // Steering piston fault closing time exceeded
         SPFopen_MH : Bool;   // Steering piston fault MH is open before shot
         SPFclosed_MH : Bool;   // Steering piston MH closed before end of shot
         MHBouncing : Bool;   // Partner has shot enabled
         SPFaborted_SoftwareRelease : Bool;
         SPFaborted_CP : Bool;
         SPFabortet_HardwareRelease : Bool;
      END_STRUCT;
      IN_Reset_Fault : Bool;
      IN_CheckMH_Shot : Bool;   // Check fault mixinghead close during shot?
   END_VAR
   VAR_IN_OUT
      IO_Any_ShotCycleState : ANY;
      IO_Any_MH_Fault : ANY;
      IO_FaultLevel1 : Bool;
      IO_FaultLevel2 : Bool;
      IO_FaultLevel3 : Bool;
      IO_NewFault : Bool;
   END_VAR
   VAR_TEMP
      Temp_Any_ShotCycleState : ANY;
      Temp_Any_MH_Fault : ANY;
      Temp_MH_Fault : "UDT1842_FLT_MH_Control";
      Tenp_ShotCycleState : "UDT091_PouringCycleState";
      ERROR_CODE : Int;
   END_VAR
BEGIN

REGION Network 1: Get temporary variables shot cycle
         L;
         LAR1;
         LAR2;
   //
         L     W[AR1, P#0.0];  // Bytes
         T     W[AR2, P#0.0];
         L     W[AR1, P#2.0];  //Amount of bytes
         T     W[AR2, P#2.0];
         L     W[AR1, P#4.0];  //Block no,
         T     W[AR2, P#4.0];
         L     D[AR1, P#6.0];  // Startadress of data
         T     D[AR2, P#6.0];
   //
         CALL  BLKMOV
         ( SRCBLK  := #Temp_Any_ShotCycleState,
           RET_VAL := #ERROR_CODE,
           DSTBLK  := #Tenp_ShotCycleState
         );
END_REGION

REGION Network 2: Get temporary variables MH fault
         L;
         LAR1;
         LAR2;
   //
         L     W[AR1, P#0.0];  // Bytes
         T     W[AR2, P#0.0];
         L     W[AR1, P#2.0];  //Amount of bytes
         T     W[AR2, P#2.0];
         L     W[AR1, P#4.0];  //Block no,
         T     W[AR2, P#4.0];
         L     D[AR1, P#6.0];  // Startadress of data
         T     D[AR2, P#6.0];
   //
         CALL  BLKMOV
         ( SRCBLK  := #Temp_Any_MH_Fault,
           RET_VAL := #ERROR_CODE,
           DSTBLK  := #Temp_MH_Fault
         );
END_REGION

REGION Network 3: Reset faults mixing head
         AN    #IN_Reset_Fault;
         JC    nw3e;

         CLR;
         =     #Temp_MH_Fault.FLT_MH_dontOpen;
         =     #Temp_MH_Fault.FLT_MH_dontClose;
         =     #Temp_MH_Fault.FLT_ShotStopped;
         =     #Temp_MH_Fault.FLT_MH_OpenWOactivation;
         =     #Temp_MH_Fault.FLT_MH_CloseDuringShot;
         =     #Temp_MH_Fault.WRN_ShotTimeShort;
         =     #Temp_MH_Fault.WRN_ShotTimeLong;
         =     #Temp_MH_Fault.FLT_ShotTimeShort;
         =     #Temp_MH_Fault.FLT_MH_bounce;

   nw3e: NOP   0;
END_REGION

REGION Network 4: Fault mixinghead from ProCan mixinghead state
         A     #IN_ProCanMH_State.SPFopening_MH;
         AN    #Temp_MH_Fault.FLT_MH_dontOpen;
         S     #Temp_MH_Fault.FLT_MH_dontOpen;
         S     #IO_NewFault;

         A     #IN_ProCanMH_State.SPFclosing_MH;
         AN    #Temp_MH_Fault.FLT_MH_dontClose;
         S     #Temp_MH_Fault.FLT_MH_dontClose;
         S     #IO_NewFault;

         O     #IN_ProCanMH_State.SPFaborted_SoftwareRelease;
         O     #IN_ProCanMH_State.SPFaborted_CP;
         O     #IN_ProCanMH_State.SPFabortet_HardwareRelease;
         AN    #Temp_MH_Fault.FLT_ShotStopped;
         S     #Temp_MH_Fault.FLT_ShotStopped;
         S     #IO_NewFault;

         A     #IN_ProCanMH_State.SPFopen_MH;
         AN    #Temp_MH_Fault.FLT_MH_OpenWOactivation;
         S     #Temp_MH_Fault.FLT_MH_OpenWOactivation;
         S     #IO_NewFault;

         A     #IN_ProCanMH_State.SPFclosed_MH;
         AN    #Temp_MH_Fault.FLT_MH_CloseDuringShot;
         S     #Temp_MH_Fault.FLT_MH_CloseDuringShot;
         S     #IO_NewFault;
END_REGION

REGION Network 5: Fault levels
         O     #Temp_MH_Fault.FLT_MH_dontOpen;
         O     #Temp_MH_Fault.FLT_MH_dontClose;
         O     #Temp_MH_Fault.FLT_MH_OpenWOactivation;
         O     #Temp_MH_Fault.FLT_MH_CloseDuringShot;
         S     #IO_FaultLevel1;

         O     #Temp_MH_Fault.FLT_ShotStopped;
         S     #IO_FaultLevel3;
END_REGION

REGION Network 6: Write back faults
         CALL  BLKMOV
         ( SRCBLK  := #Temp_MH_Fault,
           RET_VAL := #ERROR_CODE,
           DSTBLK  := #Temp_Any_MH_Fault
         );
END_REGION
END_FUNCTION

FUNCTION "FC101_auxiliaryDrive" : Void   // FC101, STL
TITLE = Control of several auxiliary drives of a pouring machine
{ S7_Optimized_Access := 'FALSE' }
AUTHOR : KT242
FAMILY : RS_KK
NAME : Drive
VERSION : 1.5
   VAR_INPUT
      IN_Release : Bool;   // Genarelly release 0f the drive (Operation mode)
      IN_ControlVoltage : Bool;   // Signal delay activation frequency converter (protection after emergency-stop)
      IN_Reset_fault : Bool;   // Signal to quit fault within function block
      IN_Request_Filling : Bool;   // Request switch on drive for filling
      IN_Request_Feedpump : Bool;   // Request switch on drive if componenten pump start up
      IN_Request_Cooling : Bool;   // Request switch on drive for cooling // runs without pause
      IN_Request_Heating : Bool;   // Request switch on drive for heating // runs with pause
      IN_Fault_Motorprotection : Bool;   // Input fault motorprotection of drive
      IN_FaultFreqConverter : Bool;   // Input fault frequency converter of drive
      IN_MaxPressure_MaxLTray : Bool;   // Input fault max. pressure or max. filling level tray
      IN_DryRun : Bool;   // Input fault Min_Level or dry run
      IN_DW_RunTime : S5Time;   // Time value of runtime of drive
      IN_DW_PauseTime : S5Time;   // Time value of pausetime of drive
      IN_TimerDrive : Timer;   // Timer of general timing of the drive
      IN_TimerStartUpFConv : Timer;   // Timer of delay start up frequency converter
      IN_Configparameter : Byte;   // Configuration: 0=normal,1=filling,2=feeding,3=Edgefilter,4=FConvert
      IN_SelectFaultLevel : Bool;   // Configuration: 0=FaultLevel3, 1=Faultlevel1
   END_VAR
   VAR_OUTPUT
      OUT_MainsContactor : Bool;   // Ouput mainscontactor drive or frequency converter
      OUT_Release_FConverter : Bool;   // Output release of frequncy converter to control rotation speed
   END_VAR
   VAR_IN_OUT
      IO_Status : ANY;   // Stores the state of the drive
      IO_NewFault : Bool;
      IO_FaultLevel_1 : Bool;
      IO_FaultLevel_3 : Bool;
      IO_Faults : ANY;
   END_VAR
   VAR_TEMP
      TEMP0 : Bool;
      Temp_IO_Status : "UDT101_auxiDriveState";   // Temporary state of drive for internal use at the program block
      ERROR_CODE : Int;   // Error state of systemfunction "BLKMOV" Blockmove
      Anyzeiger1 : ANY;   // Pointer to copy thr array "IO_Status" and "Temp_IO_Status"
      Anyzeiger2 : ANY;   // Pointer to copy thr array "IO_Status" and "Temp_IO_Status"
      Temp_RunTime : S5Time;   // Flag runtime drive
      Temp_PauseTime : S5Time;   // Flag pause time
      Temp_Runtime_ms : Time;   // Flag runtime drive in millisecond
      Temp_Pausetime_ms : Time;   // Flag pause time drive in millisecond
      Temp_ReleaseDrive : Bool;   // Flag release activation drive
      Temp_IO_Fault : "UDT1801_FLT_auxDrive";
      Temp_Fault_Drive : Bool;
      Temp_MainsContactor : Bool;
      Temp_Release_FConverter : Bool;
   END_VAR
BEGIN

REGION Network 1: Saved data integration
   // Änderungen:
   // -------------------------------------------------------------------------------
   // Bei der Verwendung der Umwälzpumpe als Speisepumpe wurde dieses bei Min. 
   // Füllstand ausgeshaltet, auch wenn dies im Zyklus auftrat. Hierdurch wurden dann 
   // auch die Materialpumpen abgeschaltet.
   // v.d.Geest     25.02.2003
   // -------------------------------------------------------------------------------
   // Bei einer Ansteuerung mit Frequenzumrichter wurde nicht auf die 
   // Störungsauswertung des Umrichters gewartet bevor die Freigabe gegeben wurde. 
   // Hierdurch kam es zu Störungen bei jedem einschalten des Aggregates.
   // A. Jäger      21.11.2003
         LAR1;
         L;
         LAR2;
   //
         L     W[AR2, P#0.0];  // Bytes
         T     W[AR1, P#0.0];
         L     W[AR2, P#2.0];  //Amount of bytes
         T     W[AR1, P#2.0];
         L     W[AR2, P#4.0];  //Block no,
         T     W[AR1, P#4.0];
         L     D[AR2, P#6.0];  //Startadress of datas
         T     D[AR1, P#6.0];
   //
         CALL  BLKMOV
         ( SRCBLK  := #Anyzeiger1,
           RET_VAL := #ERROR_CODE,
           DSTBLK  := #Temp_IO_Status
         );
   //

         LAR1;
         L;
         LAR2;
   //
         L     W[AR2, P#0.0];  // Bytes
         T     W[AR1, P#0.0];
         L     W[AR2, P#2.0];  //Amount of bytes
         T     W[AR1, P#2.0];
         L     W[AR2, P#4.0];  //Block no,
         T     W[AR1, P#4.0];
         L     D[AR2, P#6.0];  //Startadress of datas
         T     D[AR1, P#6.0];
   //
         CALL  BLKMOV
         ( SRCBLK  := #Anyzeiger2,
           RET_VAL := #ERROR_CODE,
           DSTBLK  := #Temp_IO_Fault
         );
   //
END_REGION

REGION Network 2: Select operation mode
   // Mit Konfigparameter kann das unterschiedliche Verhalten eingestellt werden.
   // 0=normal      (Rührwerk,Wärmetauscher,Umwälzpumpe normal)
   // 1=charging    (Umwälzpumpe ist zugleich Befüllpumpe)
   // 2=feeding     (Umwälzpumpe ist zugleich Speisepumpe)
   // 3=edgefilter  (Splitfilter - Spaltfilter)
   // 4=fconvert    (mit FU z.B. für Rührwerk)
   // 
   // 
   // Ab Version 2.6 ist Konfigparameter nur noch ein byte, damit kompatibel zu MP270 
   // und OP's!
         SET;
         R     #Temp_IO_Status.Config_bit_normal;
         R     #Temp_IO_Status.Config_bit_char;
         R     #Temp_IO_Status.config_bit_feed;
         R     #Temp_IO_Status.Config_bit_split;  // edgefilter
         R     #Temp_IO_Status.Config_bit_with_FC;
   //
         L     #IN_Configparameter;
         JL    norm;  // case n
         JU    norm;  // case 0
         JU    char;  // case 1
         JU    feed;  // case 2
         JU    spli;  // case 3
         JU    fu;  // case 4
   norm: SET;
         =     #Temp_IO_Status.Config_bit_normal;
         JU    end;
   char: SET;
         =     #Temp_IO_Status.Config_bit_char;
         JU    end;
   feed: SET;
         =     #Temp_IO_Status.config_bit_feed;
         JU    end;
   spli: SET;
         =     #Temp_IO_Status.Config_bit_split;
         JU    end;
   fu:   SET;
         =     #Temp_IO_Status.Config_bit_with_FC;
   end:  NOP   0;
END_REGION

